REGION Network 8: Concatenadora 2
   RUNG wire#powerrail
      Contact( "EstadosCmpALTA-MTA"._5s4 )
      wire#w1
      { S7_Templates := "SrcType := Int" } NE_Contact(in1 := "CompALTA-MTA".VRealCmp5, in2 := 1)
      wire#w2
      { S7_Templates := "SrcType := Int" } GT_Contact(in1 := "CompALTA-MTA".VRealCmp5, in2 := "CompALTA-MTA".VRealCmp1)
      { S7_Templates := "SrcType := Int" } NE_Contact(in1 := "CompALTA-MTA".VRealCmp1, in2 := 0)
      wire#w3
      Contact( "TV5" )
      wire#w4
      Coil( "Concatenadoras"._5c2 )
   END_RUNG
   RUNG wire#w2
      { S7_Templates := "SrcType := Int" } GT_Contact(in1 := "CompALTA-MTA".VRealCmp5, in2 := "CompALTA-MTA".VRealCmp2)
      { S7_Templates := "SrcType := Int" } NE_Contact(in1 := "CompALTA-MTA".VRealCmp2, in2 := 0)
   END_RUNG wire#w3
   RUNG wire#w2
      { S7_Templates := "SrcType := Int" } GT_Contact(in1 := "CompALTA-MTA".VRealCmp5, in2 := "CompALTA-MTA".VRealCmp3)
      { S7_Templates := "SrcType := Int" } NE_Contact(in1 := "CompALTA-MTA".VRealCmp3, in2 := 0)
   END_RUNG wire#w3
   RUNG wire#w2
      { S7_Templates := "SrcType := Int" } GT_Contact(in1 := "CompALTA-MTA".VRealCmp5, in2 := "CompALTA-MTA".VRealCmp4)
      { S7_Templates := "SrcType := Int" } NE_Contact(in1 := "CompALTA-MTA".VRealCmp4, in2 := 0)
   END_RUNG wire#w3
   RUNG wire#w2
      { S7_Templates := "SrcType := Int" } GT_Contact(in1 := "CompALTA-MTA".VRealCmp5, in2 := "CompALTA-MTA".VRealCmp6)
      { S7_Templates := "SrcType := Int" } NE_Contact(in1 := "CompALTA-MTA".VRealCmp6, in2 := 0)
   END_RUNG wire#w3
   RUNG wire#w1
      Contact( "DB-CompAltaDatos".TON_ParGenMem )
   END_RUNG wire#w4
   RUNG wire#powerrail
      Contact( "EstadosCmpALTA-MTA"._5s6 )
      Contact( "DB-CompAltaDatos".Aut5 )
      Contact( "DB-CompAltaDatos".PanMchCmp5 )
   END_RUNG wire#w4
   // the same network as SCL:
   "Concatenadoras"._5c2 := ("EstadosCmpALTA-MTA"._5s4 AND ((("CompALTA-MTA".VRealCmp5 <> 1) AND ((("CompALTA-MTA".VRealCmp5 > "CompALTA-MTA".VRealCmp1) AND ("CompALTA-MTA".VRealCmp1 <> 0)) OR (("CompALTA-MTA".VRealCmp5 > "CompALTA-MTA".VRealCmp2) AND ("CompALTA-MTA".VRealCmp2 <> 0)) OR (("CompALTA-MTA".VRealCmp5 > "CompALTA-MTA".VRealCmp3) AND ("CompALTA-MTA".VRealCmp3 <> 0)) OR (("CompALTA-MTA".VRealCmp5 > "CompALTA-MTA".VRealCmp4) AND ("CompALTA-MTA".VRealCmp4 <> 0)) OR (("CompALTA-MTA".VRealCmp5 > "CompALTA-MTA".VRealCmp6) AND ("CompALTA-MTA".VRealCmp6 <> 0))) AND "TV5") OR "DB-CompAltaDatos".TON_ParGenMem)) OR ("EstadosCmpALTA-MTA"._5s6 AND "DB-CompAltaDatos".Aut5 AND "DB-CompAltaDatos".PanMchCmp5);
END_REGION

REGION Network 9: Concatenadora 3
   RUNG wire#powerrail
      Contact( "EstadosCmpALTA-MTA"._5s2 )
      Contact( "TsinReq5" )
      wire#w1
      Coil( "Concatenadoras"._5c3 )
   END_RUNG
   RUNG wire#powerrail
      Contact( "EstadosCmpALTA-MTA"._5s10 )
      Contact( "DB-CompAltaDatos".PanMchCmp5 )
   END_RUNG wire#w1
   // the same network as SCL:
   "Concatenadoras"._5c3 := ("EstadosCmpALTA-MTA"._5s2 AND "TsinReq5") OR ("EstadosCmpALTA-MTA"._5s10 AND "DB-CompAltaDatos".PanMchCmp5);
END_REGION

REGION Network 10: Concatenadora 10
   RUNG wire#powerrail
      Contact( "EstadosCmpALTA-MTA"._5s1 )
      I_Contact( "CompALTA-MTA".ReqMch5 )
      wire#w1
      Contact( "DB-CompAltaDatos".Aut5 )
      Coil( "Concatenadoras"._5c10 )
   END_RUNG
   RUNG wire#powerrail
      Contact( "EstadosCmpALTA-MTA"._5s9 )
      I_Contact( "CompALTA-MTA".ReqMch5 )
   END_RUNG wire#w1
   RUNG wire#powerrail
      Contact( "EstadosCmpALTA-MTA"._5s3 )
      I_Contact( "DB-CompAltaDatos".PanMchCmp5 )
   END_RUNG wire#w1
   // the same network as SCL:
   "Concatenadoras"._5c10 := (("EstadosCmpALTA-MTA"._5s1 AND NOT "CompALTA-MTA".ReqMch5) OR ("EstadosCmpALTA-MTA"._5s9 AND NOT "CompALTA-MTA".ReqMch5) OR ("EstadosCmpALTA-MTA"._5s3 AND NOT "DB-CompAltaDatos".PanMchCmp5)) AND "DB-CompAltaDatos".Aut5;
END_REGION

REGION Network 11: Concatenadora 4
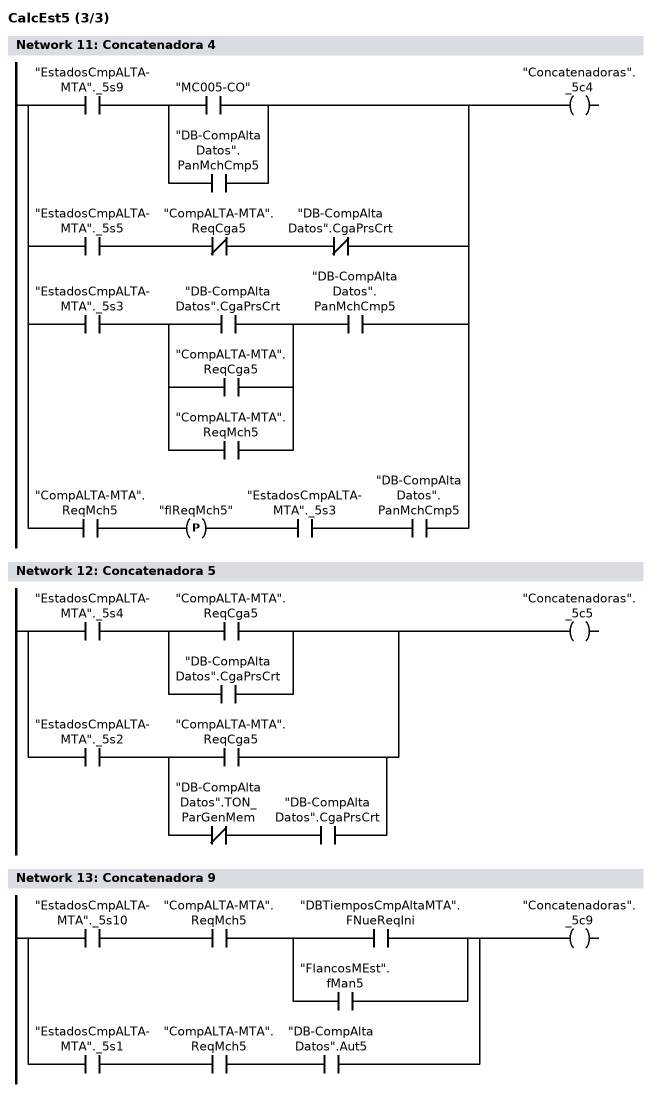
   RUNG wire#powerrail
      Contact( "EstadosCmpALTA-MTA"._5s9 )
      wire#w1
      Contact( "MC005-CO" )
      wire#w2
      Coil( "Concatenadoras"._5c4 )
   END_RUNG
   RUNG wire#w1
      Contact( "DB-CompAltaDatos".PanMchCmp5 )
   END_RUNG wire#w2
   RUNG wire#powerrail
      Contact( "EstadosCmpALTA-MTA"._5s5 )
      I_Contact( "CompALTA-MTA".ReqCga5 )
      I_Contact( "DB-CompAltaDatos".CgaPrsCrt )
   END_RUNG wire#w2
   RUNG wire#powerrail
      Contact( "EstadosCmpALTA-MTA"._5s3 )
      wire#w3
      Contact( "DB-CompAltaDatos".CgaPrsCrt )
      wire#w4
      Contact( "DB-CompAltaDatos".PanMchCmp5 )
   END_RUNG wire#w2
   RUNG wire#w3
      Contact( "CompALTA-MTA".ReqCga5 )
   END_RUNG wire#w4
   RUNG wire#w3
      Contact( "CompALTA-MTA".ReqMch5 )
   END_RUNG wire#w4
   RUNG wire#powerrail
      Contact( "CompALTA-MTA".ReqMch5 )
      P_Trig( "flReqMch5" )
      Contact( "EstadosCmpALTA-MTA"._5s3 )
      Contact( "DB-CompAltaDatos".PanMchCmp5 )
   END_RUNG wire#w2
   // the same network as SCL:
   #_w1 := "CompALTA-MTA".ReqMch5 AND NOT "flReqMch5";   // rising edge
   "flReqMch5" := "CompALTA-MTA".ReqMch5;
   "Concatenadoras"._5c4 := ("EstadosCmpALTA-MTA"._5s9 AND ("MC005-CO" OR "DB-CompAltaDatos".PanMchCmp5)) OR ("EstadosCmpALTA-MTA"._5s5 AND NOT "CompALTA-MTA".ReqCga5 AND NOT "DB-CompAltaDatos".CgaPrsCrt) OR ("EstadosCmpALTA-MTA"._5s3 AND ("DB-CompAltaDatos".CgaPrsCrt OR "CompALTA-MTA".ReqCga5 OR "CompALTA-MTA".ReqMch5) AND "DB-CompAltaDatos".PanMchCmp5) OR (#_w1 AND "EstadosCmpALTA-MTA"._5s3 AND "DB-CompAltaDatos".PanMchCmp5);
END_REGION

REGION Network 12: Concatenadora 5
   RUNG wire#powerrail
      Contact( "EstadosCmpALTA-MTA"._5s4 )
      wire#w1
      Contact( "CompALTA-MTA".ReqCga5 )
      wire#w2
      Coil( "Concatenadoras"._5c5 )
   END_RUNG
   RUNG wire#w1
      Contact( "DB-CompAltaDatos".CgaPrsCrt )
   END_RUNG wire#w2
   RUNG wire#powerrail
      Contact( "EstadosCmpALTA-MTA"._5s2 )
      wire#w3
      Contact( "CompALTA-MTA".ReqCga5 )
   END_RUNG wire#w2
   RUNG wire#w3
      I_Contact( "DB-CompAltaDatos".TON_ParGenMem )
      Contact( "DB-CompAltaDatos".CgaPrsCrt )
   END_RUNG wire#w2
   // the same network as SCL:
   "Concatenadoras"._5c5 := ("EstadosCmpALTA-MTA"._5s4 AND ("CompALTA-MTA".ReqCga5 OR "DB-CompAltaDatos".CgaPrsCrt)) OR ("EstadosCmpALTA-MTA"._5s2 AND ("CompALTA-MTA".ReqCga5 OR (NOT "DB-CompAltaDatos".TON_ParGenMem AND "DB-CompAltaDatos".CgaPrsCrt)));
END_REGION

REGION Network 13: Concatenadora 9
   RUNG wire#powerrail
      Contact( "EstadosCmpALTA-MTA"._5s10 )
      Contact( "CompALTA-MTA".ReqMch5 )
      wire#w1
      Contact( "DBTiemposCmpAltaMTA".FNueReqIni )
      wire#w2
      Coil( "Concatenadoras"._5c9 )
   END_RUNG
   RUNG wire#w1
      Contact( "FlancosMEst".fMan5 )
   END_RUNG wire#w2
   RUNG wire#powerrail
      Contact( "EstadosCmpALTA-MTA"._5s1 )
      Contact( "CompALTA-MTA".ReqMch5 )
      Contact( "DB-CompAltaDatos".Aut5 )
   END_RUNG wire#w2
   // the same network as SCL:
   "Concatenadoras"._5c9 := ("EstadosCmpALTA-MTA"._5s10 AND "CompALTA-MTA".ReqMch5 AND ("DBTiemposCmpAltaMTA".FNueReqIni OR "FlancosMEst".fMan5)) OR ("EstadosCmpALTA-MTA"._5s1 AND "CompALTA-MTA".ReqMch5 AND "DB-CompAltaDatos".Aut5);
END_REGION

REGION Network 14 (STL): Maquina de estados
         CALL  "FC_MAQ_EST_16"
         ( IN0  := %DB127.DBW8,
           IN1  := %DB128.DBW8,
           OUT2 := "ErrPMQ5",
           OUT3 := "ErrCMQ5",
           IO4  := %DB120.DBW8
         );
         NOP   0;
END_REGION

REGION Network 15 (STL): Bloque animación compresor
         CALL  "FC-ANIM-CMP"
         ( IN0  := %DB120.DBW8,
           OUT1 := "CompALTA-MTA".AnimCMP5
         );
         NOP   0;
END_REGION
END_FUNCTION

FUNCTION "CalcEst0" : Void   // FC42, LAD
{ S7_Optimized_Access := 'FALSE' }
VERSION : 0.1
BEGIN

REGION Network 1
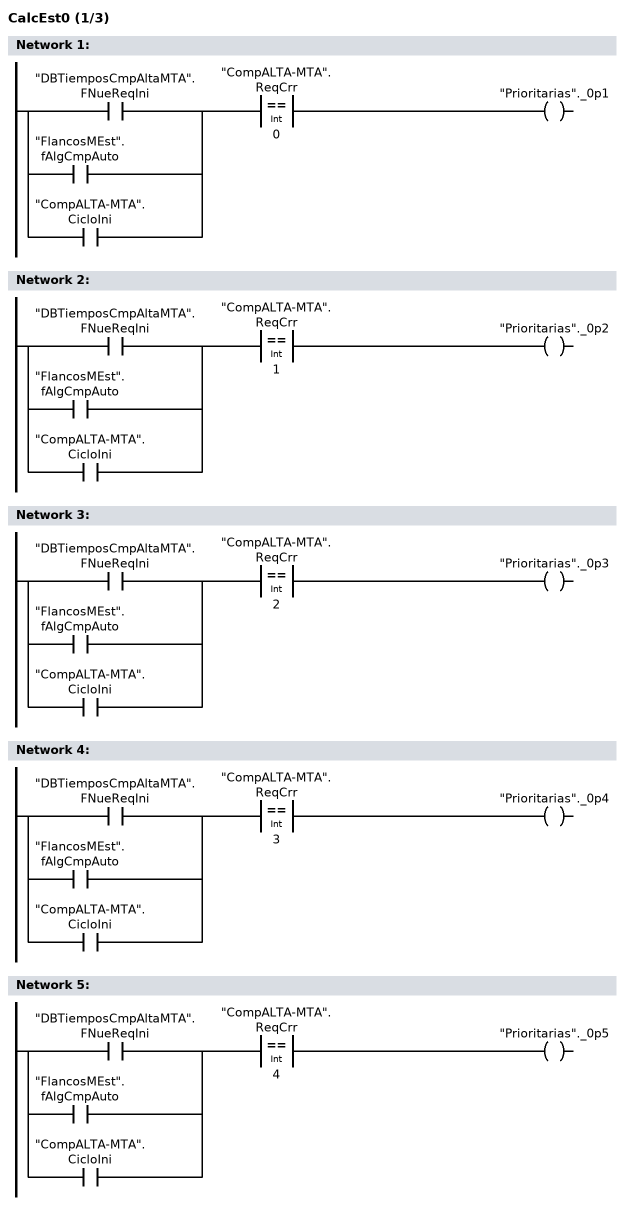
   RUNG wire#powerrail
      Contact( "DBTiemposCmpAltaMTA".FNueReqIni )
      wire#w1
      { S7_Templates := "SrcType := Int" } EQ_Contact(in1 := "CompALTA-MTA".ReqCrr, in2 := 0)
      Coil( "Prioritarias"._0p1 )
   END_RUNG
   RUNG wire#powerrail
      Contact( "FlancosMEst".fAlgCmpAuto )
   END_RUNG wire#w1
   RUNG wire#powerrail
      Contact( "CompALTA-MTA".CicloIni )
   END_RUNG wire#w1
   // the same network as SCL:
   "Prioritarias"._0p1 := ("DBTiemposCmpAltaMTA".FNueReqIni OR "FlancosMEst".fAlgCmpAuto OR "CompALTA-MTA".CicloIni) AND ("CompALTA-MTA".ReqCrr = 0);
END_REGION

REGION Network 2
   RUNG wire#powerrail
      Contact( "DBTiemposCmpAltaMTA".FNueReqIni )
      wire#w1
      { S7_Templates := "SrcType := Int" } EQ_Contact(in1 := "CompALTA-MTA".ReqCrr, in2 := 1)
      Coil( "Prioritarias"._0p2 )
   END_RUNG
   RUNG wire#powerrail
      Contact( "FlancosMEst".fAlgCmpAuto )
   END_RUNG wire#w1
   RUNG wire#powerrail
      Contact( "CompALTA-MTA".CicloIni )
   END_RUNG wire#w1
   // the same network as SCL:
   "Prioritarias"._0p2 := ("DBTiemposCmpAltaMTA".FNueReqIni OR "FlancosMEst".fAlgCmpAuto OR "CompALTA-MTA".CicloIni) AND ("CompALTA-MTA".ReqCrr = 1);
END_REGION

REGION Network 3
   RUNG wire#powerrail
      Contact( "DBTiemposCmpAltaMTA".FNueReqIni )
      wire#w1
      { S7_Templates := "SrcType := Int" } EQ_Contact(in1 := "CompALTA-MTA".ReqCrr, in2 := 2)
      Coil( "Prioritarias"._0p3 )
   END_RUNG
   RUNG wire#powerrail
      Contact( "FlancosMEst".fAlgCmpAuto )
   END_RUNG wire#w1
   RUNG wire#powerrail
      Contact( "CompALTA-MTA".CicloIni )
   END_RUNG wire#w1
   // the same network as SCL:
   "Prioritarias"._0p3 := ("DBTiemposCmpAltaMTA".FNueReqIni OR "FlancosMEst".fAlgCmpAuto OR "CompALTA-MTA".CicloIni) AND ("CompALTA-MTA".ReqCrr = 2);
END_REGION

REGION Network 4
   RUNG wire#powerrail
      Contact( "DBTiemposCmpAltaMTA".FNueReqIni )
      wire#w1
      { S7_Templates := "SrcType := Int" } EQ_Contact(in1 := "CompALTA-MTA".ReqCrr, in2 := 3)
      Coil( "Prioritarias"._0p4 )
   END_RUNG
   RUNG wire#powerrail
      Contact( "FlancosMEst".fAlgCmpAuto )
   END_RUNG wire#w1
   RUNG wire#powerrail
      Contact( "CompALTA-MTA".CicloIni )
   END_RUNG wire#w1
   // the same network as SCL:
   "Prioritarias"._0p4 := ("DBTiemposCmpAltaMTA".FNueReqIni OR "FlancosMEst".fAlgCmpAuto OR "CompALTA-MTA".CicloIni) AND ("CompALTA-MTA".ReqCrr = 3);
END_REGION

REGION Network 5
   RUNG wire#powerrail
      Contact( "DBTiemposCmpAltaMTA".FNueReqIni )
      wire#w1
      { S7_Templates := "SrcType := Int" } EQ_Contact(in1 := "CompALTA-MTA".ReqCrr, in2 := 4)
      Coil( "Prioritarias"._0p5 )
   END_RUNG
   RUNG wire#powerrail
      Contact( "FlancosMEst".fAlgCmpAuto )
   END_RUNG wire#w1
   RUNG wire#powerrail
      Contact( "CompALTA-MTA".CicloIni )
   END_RUNG wire#w1
   // the same network as SCL:
   "Prioritarias"._0p5 := ("DBTiemposCmpAltaMTA".FNueReqIni OR "FlancosMEst".fAlgCmpAuto OR "CompALTA-MTA".CicloIni) AND ("CompALTA-MTA".ReqCrr = 4);
END_REGION

REGION Network 6
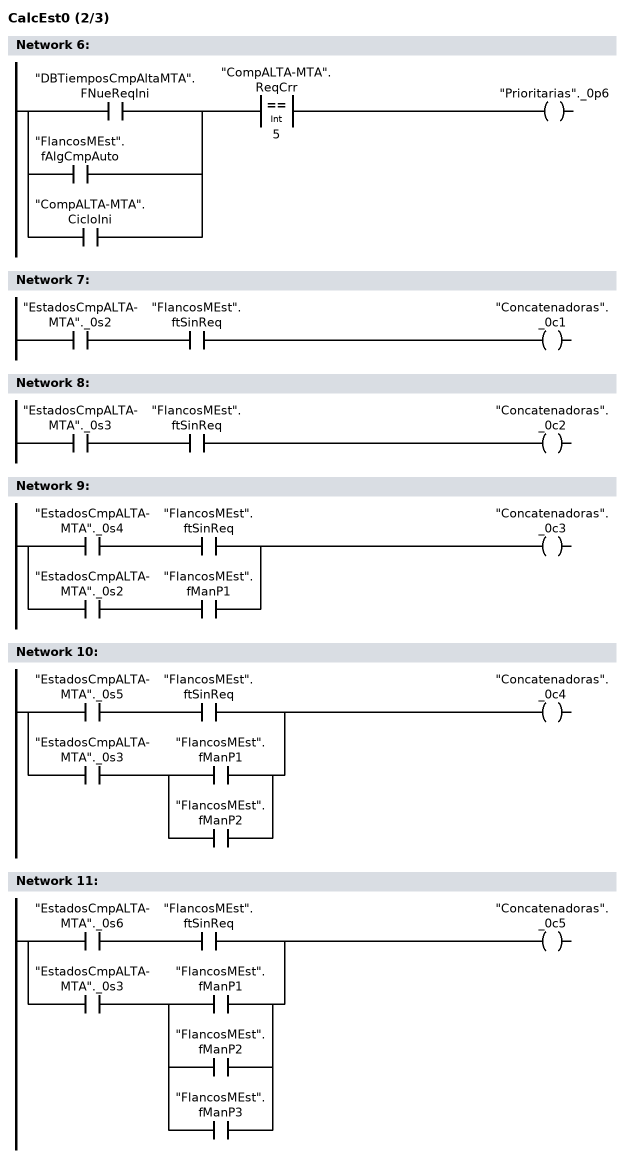
   RUNG wire#powerrail
      Contact( "DBTiemposCmpAltaMTA".FNueReqIni )
      wire#w1
      { S7_Templates := "SrcType := Int" } EQ_Contact(in1 := "CompALTA-MTA".ReqCrr, in2 := 5)
      Coil( "Prioritarias"._0p6 )
   END_RUNG
   RUNG wire#powerrail
      Contact( "FlancosMEst".fAlgCmpAuto )
   END_RUNG wire#w1
   RUNG wire#powerrail
      Contact( "CompALTA-MTA".CicloIni )
   END_RUNG wire#w1
   // the same network as SCL:
   "Prioritarias"._0p6 := ("DBTiemposCmpAltaMTA".FNueReqIni OR "FlancosMEst".fAlgCmpAuto OR "CompALTA-MTA".CicloIni) AND ("CompALTA-MTA".ReqCrr = 5);
END_REGION

REGION Network 7
   RUNG wire#powerrail
      Contact( "EstadosCmpALTA-MTA"._0s2 )
      Contact( "FlancosMEst".ftSinReq )
      Coil( "Concatenadoras"._0c1 )
   END_RUNG
   // the same network as SCL:
   "Concatenadoras"._0c1 := "EstadosCmpALTA-MTA"._0s2 AND "FlancosMEst".ftSinReq;
END_REGION

REGION Network 8
   RUNG wire#powerrail
      Contact( "EstadosCmpALTA-MTA"._0s3 )
      Contact( "FlancosMEst".ftSinReq )
      Coil( "Concatenadoras"._0c2 )
   END_RUNG
   // the same network as SCL:
   "Concatenadoras"._0c2 := "EstadosCmpALTA-MTA"._0s3 AND "FlancosMEst".ftSinReq;
END_REGION

REGION Network 9
   RUNG wire#powerrail
      Contact( "EstadosCmpALTA-MTA"._0s4 )
      Contact( "FlancosMEst".ftSinReq )
      wire#w1
      Coil( "Concatenadoras"._0c3 )
   END_RUNG
   RUNG wire#powerrail
      Contact( "EstadosCmpALTA-MTA"._0s2 )
      Contact( "FlancosMEst".fManP1 )
   END_RUNG wire#w1
   // the same network as SCL:
   "Concatenadoras"._0c3 := ("EstadosCmpALTA-MTA"._0s4 AND "FlancosMEst".ftSinReq) OR ("EstadosCmpALTA-MTA"._0s2 AND "FlancosMEst".fManP1);
END_REGION

REGION Network 10
   RUNG wire#powerrail
      Contact( "EstadosCmpALTA-MTA"._0s5 )
      Contact( "FlancosMEst".ftSinReq )
      wire#w1
      Coil( "Concatenadoras"._0c4 )
   END_RUNG
   RUNG wire#powerrail
      Contact( "EstadosCmpALTA-MTA"._0s3 )
      wire#w2
      Contact( "FlancosMEst".fManP1 )
   END_RUNG wire#w1
   RUNG wire#w2
      Contact( "FlancosMEst".fManP2 )
   END_RUNG wire#w1
   // the same network as SCL:
   "Concatenadoras"._0c4 := ("EstadosCmpALTA-MTA"._0s5 AND "FlancosMEst".ftSinReq) OR ("EstadosCmpALTA-MTA"._0s3 AND ("FlancosMEst".fManP1 OR "FlancosMEst".fManP2));
END_REGION

REGION Network 11
   RUNG wire#powerrail
      Contact( "EstadosCmpALTA-MTA"._0s6 )
      Contact( "FlancosMEst".ftSinReq )
      wire#w1
      Coil( "Concatenadoras"._0c5 )
   END_RUNG
   RUNG wire#powerrail
      Contact( "EstadosCmpALTA-MTA"._0s3 )
      wire#w2
      Contact( "FlancosMEst".fManP1 )
   END_RUNG wire#w1
   RUNG wire#w2
      Contact( "FlancosMEst".fManP2 )
   END_RUNG wire#w1
   RUNG wire#w2
      Contact( "FlancosMEst".fManP3 )
   END_RUNG wire#w1
   // the same network as SCL:
   "Concatenadoras"._0c5 := ("EstadosCmpALTA-MTA"._0s6 AND "FlancosMEst".ftSinReq) OR ("EstadosCmpALTA-MTA"._0s3 AND ("FlancosMEst".fManP1 OR "FlancosMEst".fManP2 OR "FlancosMEst".fManP3));
END_REGION

REGION Network 12
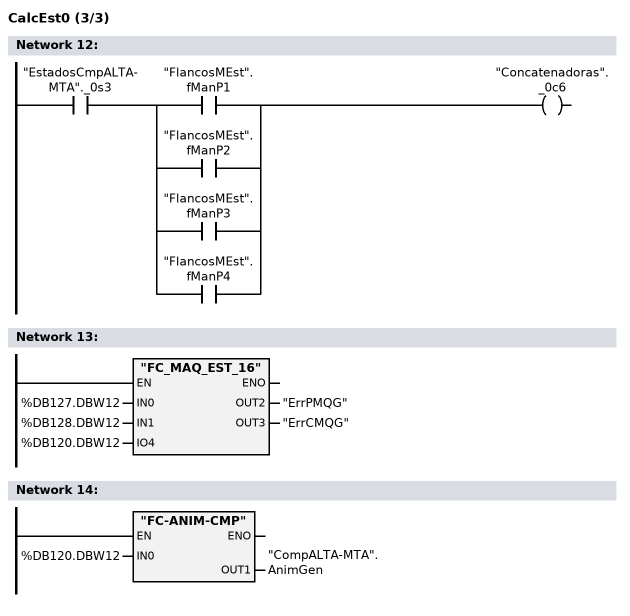
   RUNG wire#powerrail
      Contact( "EstadosCmpALTA-MTA"._0s3 )
      wire#w1
      Contact( "FlancosMEst".fManP1 )
      wire#w2
      Coil( "Concatenadoras"._0c6 )
   END_RUNG
   RUNG wire#w1
      Contact( "FlancosMEst".fManP2 )
   END_RUNG wire#w2
   RUNG wire#w1
      Contact( "FlancosMEst".fManP3 )
   END_RUNG wire#w2
   RUNG wire#w1
      Contact( "FlancosMEst".fManP4 )
   END_RUNG wire#w2
   // the same network as SCL:
   "Concatenadoras"._0c6 := "EstadosCmpALTA-MTA"._0s3 AND ("FlancosMEst".fManP1 OR "FlancosMEst".fManP2 OR "FlancosMEst".fManP3 OR "FlancosMEst".fManP4);
END_REGION

REGION Network 13
   RUNG wire#powerrail
      "FC_MAQ_EST_16"(IN0 := %DB127.DBW12, IN1 := %DB128.DBW12, IO4 := %DB120.DBW12, OUT2 => "ErrPMQG", OUT3 => "ErrCMQG")
   END_RUNG
   // the same network as SCL:
   "FC_MAQ_EST_16"(IN0 := %DB127.DBW12,
                   IN1 := %DB128.DBW12,
                   IO4 := %DB120.DBW12,
                   OUT2 => "ErrPMQG",
                   OUT3 => "ErrCMQG");
END_REGION

REGION Network 14
   RUNG wire#powerrail
      "FC-ANIM-CMP"(IN0 := %DB120.DBW12, OUT1 => "CompALTA-MTA".AnimGen)
   END_RUNG
   // the same network as SCL:
   "FC-ANIM-CMP"(IN0 := %DB120.DBW12, OUT1 => "CompALTA-MTA".AnimGen);
END_REGION
END_FUNCTION

FUNCTION "CorreccReqCmpAlta" : Void   // FC44, LAD
{ S7_Optimized_Access := 'FALSE' }
VERSION : 0.1
BEGIN

REGION Network 1
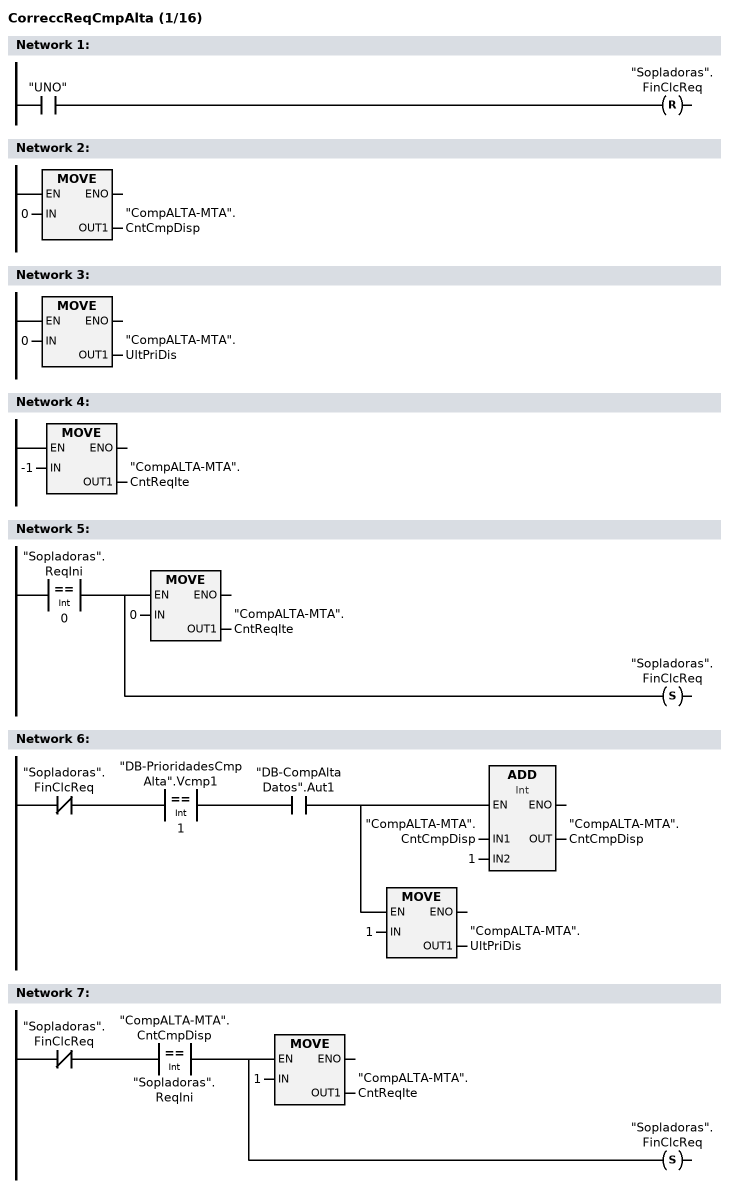
   RUNG wire#powerrail
      Contact( "UNO" )
      R_Coil( "Sopladoras".FinClcReq )
   END_RUNG
   // the same network as SCL:
   IF "UNO" THEN "Sopladoras".FinClcReq := FALSE; END_IF;
END_REGION

REGION Network 2
   RUNG wire#powerrail
      { S7_GenerateENO := "TRUE" } Move(in := 0, out1 => "CompALTA-MTA".CntCmpDisp)
   END_RUNG
   // the same network as SCL:
   "CompALTA-MTA".CntCmpDisp := 0;
END_REGION

REGION Network 3
   RUNG wire#powerrail
      { S7_GenerateENO := "TRUE" } Move(in := 0, out1 => "CompALTA-MTA".UltPriDis)
   END_RUNG
   // the same network as SCL:
   "CompALTA-MTA".UltPriDis := 0;
END_REGION

REGION Network 4
   RUNG wire#powerrail
      { S7_GenerateENO := "TRUE" } Move(in := -1, out1 => "CompALTA-MTA".CntReqIte)
   END_RUNG
   // the same network as SCL:
   "CompALTA-MTA".CntReqIte := -1;
END_REGION

REGION Network 5
   RUNG wire#powerrail
      { S7_Templates := "SrcType := Int" } EQ_Contact(in1 := "Sopladoras".ReqIni, in2 := 0)
      wire#w1
      { S7_GenerateENO := "TRUE" } Move(in := 0, out1 => "CompALTA-MTA".CntReqIte)
   END_RUNG
   RUNG wire#w1
      S_Coil( "Sopladoras".FinClcReq )
   END_RUNG
   // the same network as SCL:
   IF "Sopladoras".ReqIni = 0 THEN
       "CompALTA-MTA".CntReqIte := 0;
       "Sopladoras".FinClcReq := TRUE;
   END_IF;
END_REGION

REGION Network 6
   IF NOT "Sopladoras".FinClcReq AND ("DB-PrioridadesCmpAlta".Vcmp1 = 1) AND "DB-CompAltaDatos".Aut1 THEN
       "CompALTA-MTA".CntCmpDisp := "CompALTA-MTA".CntCmpDisp + 1;
       "CompALTA-MTA".UltPriDis := 1;
   END_IF;
END_REGION

REGION Network 7
   IF NOT "Sopladoras".FinClcReq AND ("CompALTA-MTA".CntCmpDisp = "Sopladoras".ReqIni) THEN
       "CompALTA-MTA".CntReqIte := 1;
       "Sopladoras".FinClcReq := TRUE;
   END_IF;
END_REGION

REGION Network 8
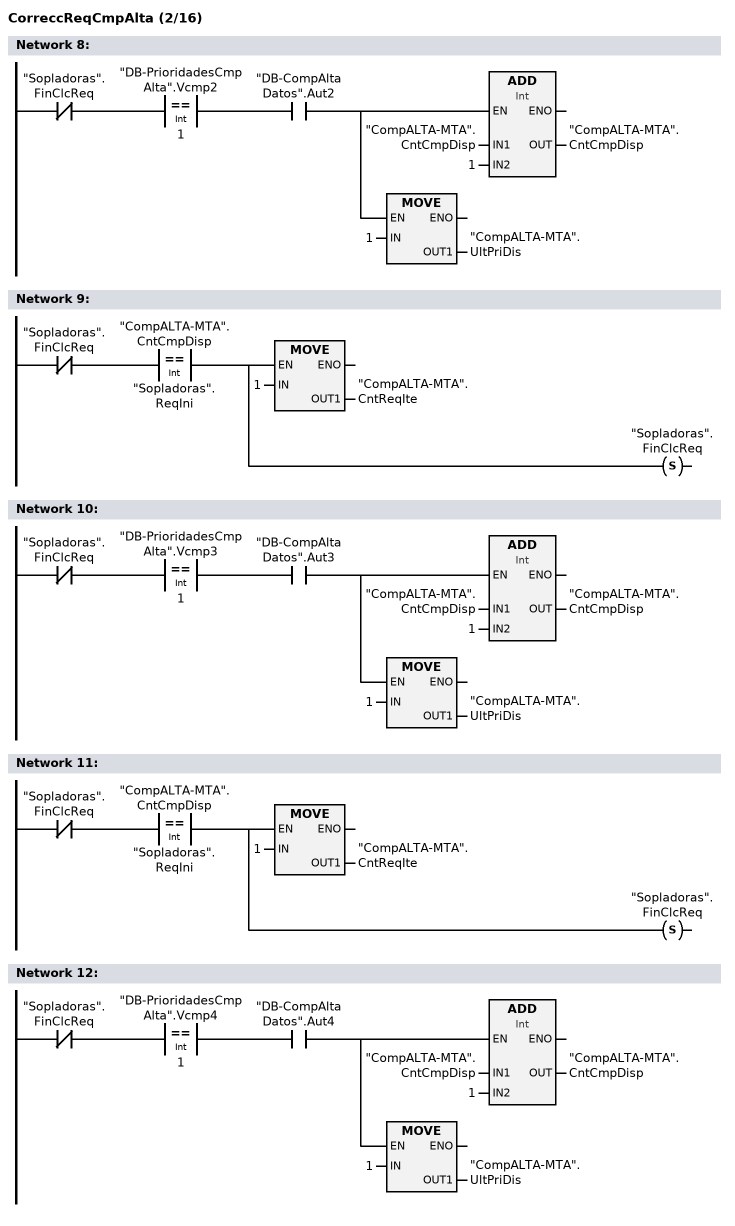
   IF NOT "Sopladoras".FinClcReq AND ("DB-PrioridadesCmpAlta".Vcmp2 = 1) AND "DB-CompAltaDatos".Aut2 THEN
       "CompALTA-MTA".CntCmpDisp := "CompALTA-MTA".CntCmpDisp + 1;
       "CompALTA-MTA".UltPriDis := 1;
   END_IF;
END_REGION

REGION Network 9
   IF NOT "Sopladoras".FinClcReq AND ("CompALTA-MTA".CntCmpDisp = "Sopladoras".ReqIni) THEN
       "CompALTA-MTA".CntReqIte := 1;
       "Sopladoras".FinClcReq := TRUE;
   END_IF;
END_REGION

REGION Network 10
   IF NOT "Sopladoras".FinClcReq AND ("DB-PrioridadesCmpAlta".Vcmp3 = 1) AND "DB-CompAltaDatos".Aut3 THEN
       "CompALTA-MTA".CntCmpDisp := "CompALTA-MTA".CntCmpDisp + 1;
       "CompALTA-MTA".UltPriDis := 1;
   END_IF;
END_REGION

REGION Network 11
   IF NOT "Sopladoras".FinClcReq AND ("CompALTA-MTA".CntCmpDisp = "Sopladoras".ReqIni) THEN
       "CompALTA-MTA".CntReqIte := 1;
       "Sopladoras".FinClcReq := TRUE;
   END_IF;
END_REGION

REGION Network 12
   IF NOT "Sopladoras".FinClcReq AND ("DB-PrioridadesCmpAlta".Vcmp4 = 1) AND "DB-CompAltaDatos".Aut4 THEN
       "CompALTA-MTA".CntCmpDisp := "CompALTA-MTA".CntCmpDisp + 1;
       "CompALTA-MTA".UltPriDis := 1;
   END_IF;
END_REGION

REGION Network 13
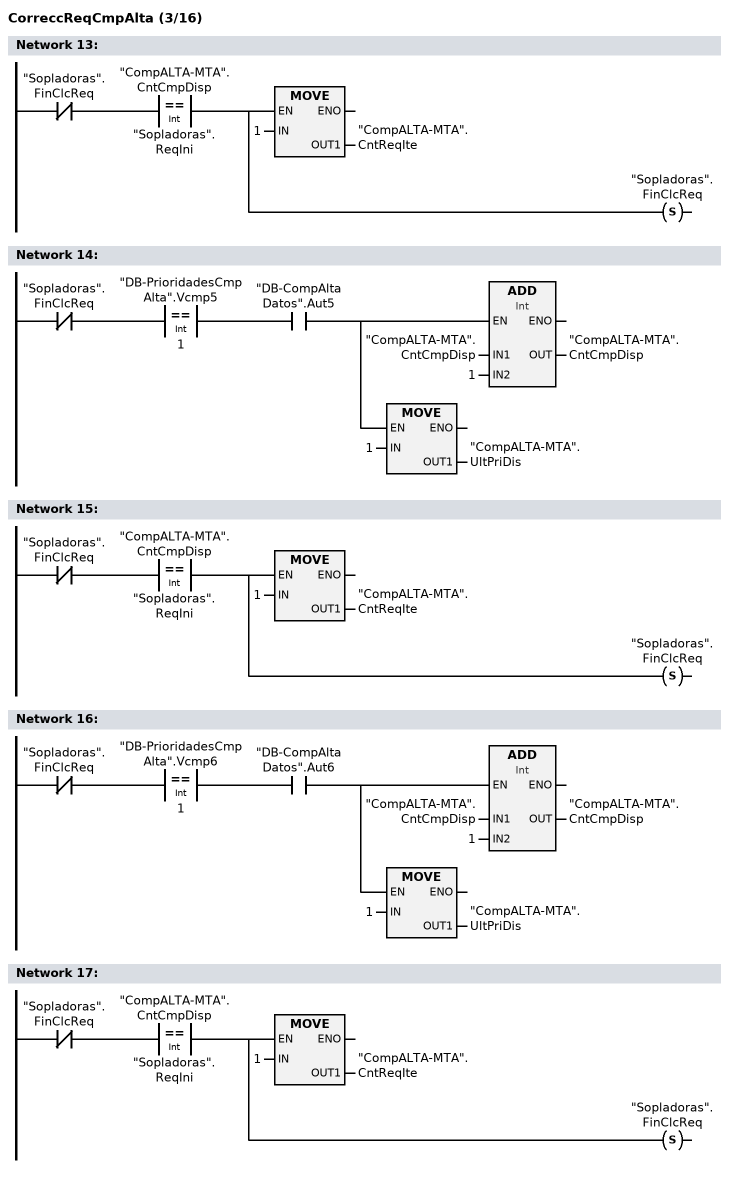
   IF NOT "Sopladoras".FinClcReq AND ("CompALTA-MTA".CntCmpDisp = "Sopladoras".ReqIni) THEN
       "CompALTA-MTA".CntReqIte := 1;
       "Sopladoras".FinClcReq := TRUE;
   END_IF;
END_REGION

REGION Network 14
   IF NOT "Sopladoras".FinClcReq AND ("DB-PrioridadesCmpAlta".Vcmp5 = 1) AND "DB-CompAltaDatos".Aut5 THEN
       "CompALTA-MTA".CntCmpDisp := "CompALTA-MTA".CntCmpDisp + 1;
       "CompALTA-MTA".UltPriDis := 1;
   END_IF;
END_REGION

REGION Network 15
   IF NOT "Sopladoras".FinClcReq AND ("CompALTA-MTA".CntCmpDisp = "Sopladoras".ReqIni) THEN
       "CompALTA-MTA".CntReqIte := 1;
       "Sopladoras".FinClcReq := TRUE;
   END_IF;
END_REGION

REGION Network 16
   RUNG wire#powerrail
      I_Contact( "Sopladoras".FinClcReq )
      { S7_Templates := "SrcType := Int" } EQ_Contact(in1 := "DB-PrioridadesCmpAlta".Vcmp6, in2 := 1)
      Contact( "DB-CompAltaDatos".Aut6 )
      wire#w1
      { S7_Templates := "SrcType := Int"; S7_GenerateENO := "TRUE" } Add(in1 := "CompALTA-MTA".CntCmpDisp, in2 := 1, out => "CompALTA-MTA".CntCmpDisp)
   END_RUNG
   RUNG wire#w1
      { S7_GenerateENO := "TRUE" } Move(in := 1, out1 => "CompALTA-MTA".UltPriDis)
   END_RUNG
   // the same network as SCL:
   IF NOT "Sopladoras".FinClcReq AND ("DB-PrioridadesCmpAlta".Vcmp6 = 1) AND "DB-CompAltaDatos".Aut6 THEN
       "CompALTA-MTA".CntCmpDisp := "CompALTA-MTA".CntCmpDisp + 1;
       "CompALTA-MTA".UltPriDis := 1;
   END_IF;
END_REGION

REGION Network 17
   RUNG wire#powerrail
      I_Contact( "Sopladoras".FinClcReq )
      { S7_Templates := "SrcType := Int" } EQ_Contact(in1 := "CompALTA-MTA".CntCmpDisp, in2 := "Sopladoras".ReqIni)
      wire#w1
      { S7_GenerateENO := "TRUE" } Move(in := 1, out1 => "CompALTA-MTA".CntReqIte)
   END_RUNG
   RUNG wire#w1
      S_Coil( "Sopladoras".FinClcReq )
   END_RUNG
   // the same network as SCL:
   IF NOT "Sopladoras".FinClcReq AND ("CompALTA-MTA".CntCmpDisp = "Sopladoras".ReqIni) THEN
       "CompALTA-MTA".CntReqIte := 1;
       "Sopladoras".FinClcReq := TRUE;
   END_IF;
END_REGION

REGION Network 18
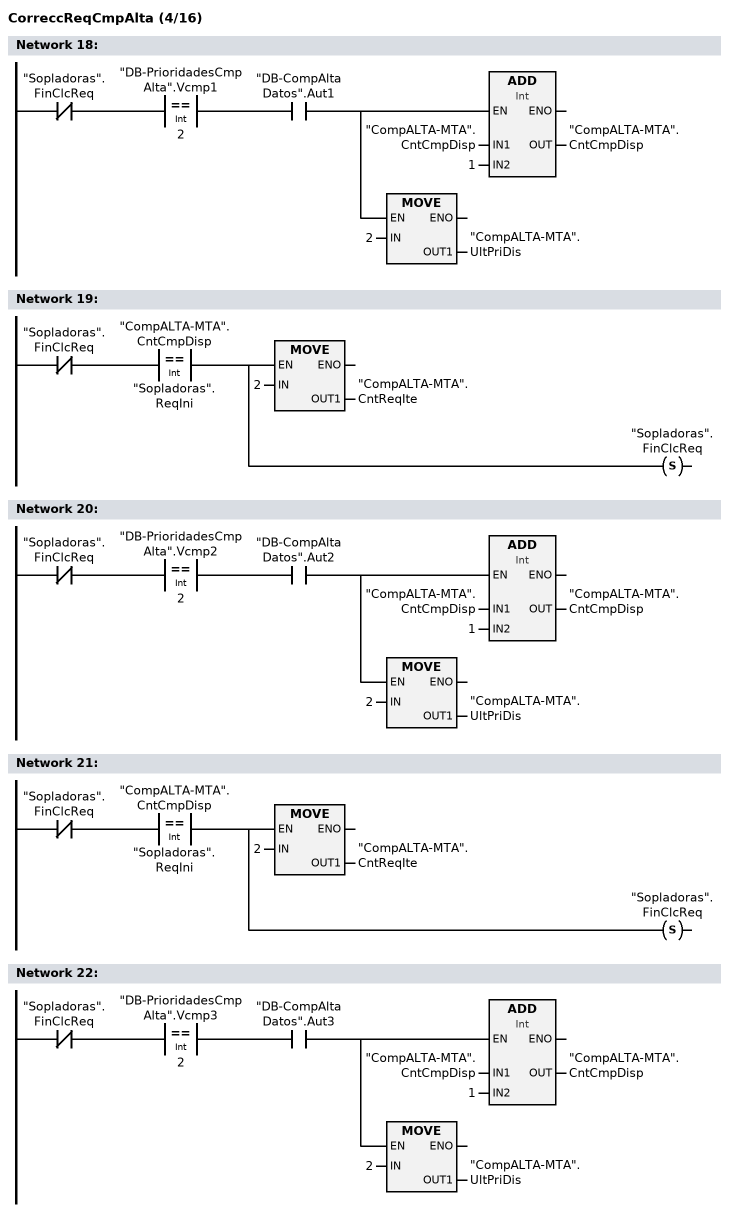
   IF NOT "Sopladoras".FinClcReq AND ("DB-PrioridadesCmpAlta".Vcmp1 = 2) AND "DB-CompAltaDatos".Aut1 THEN
       "CompALTA-MTA".CntCmpDisp := "CompALTA-MTA".CntCmpDisp + 1;
       "CompALTA-MTA".UltPriDis := 2;
   END_IF;
END_REGION

REGION Network 19
   IF NOT "Sopladoras".FinClcReq AND ("CompALTA-MTA".CntCmpDisp = "Sopladoras".ReqIni) THEN
       "CompALTA-MTA".CntReqIte := 2;
       "Sopladoras".FinClcReq := TRUE;
   END_IF;
END_REGION

REGION Network 20
   IF NOT "Sopladoras".FinClcReq AND ("DB-PrioridadesCmpAlta".Vcmp2 = 2) AND "DB-CompAltaDatos".Aut2 THEN
       "CompALTA-MTA".CntCmpDisp := "CompALTA-MTA".CntCmpDisp + 1;
       "CompALTA-MTA".UltPriDis := 2;
   END_IF;
END_REGION

REGION Network 21
   IF NOT "Sopladoras".FinClcReq AND ("CompALTA-MTA".CntCmpDisp = "Sopladoras".ReqIni) THEN
       "CompALTA-MTA".CntReqIte := 2;
       "Sopladoras".FinClcReq := TRUE;
   END_IF;
END_REGION

REGION Network 22
   IF NOT "Sopladoras".FinClcReq AND ("DB-PrioridadesCmpAlta".Vcmp3 = 2) AND "DB-CompAltaDatos".Aut3 THEN
       "CompALTA-MTA".CntCmpDisp := "CompALTA-MTA".CntCmpDisp + 1;
       "CompALTA-MTA".UltPriDis := 2;
   END_IF;
END_REGION

REGION Network 23
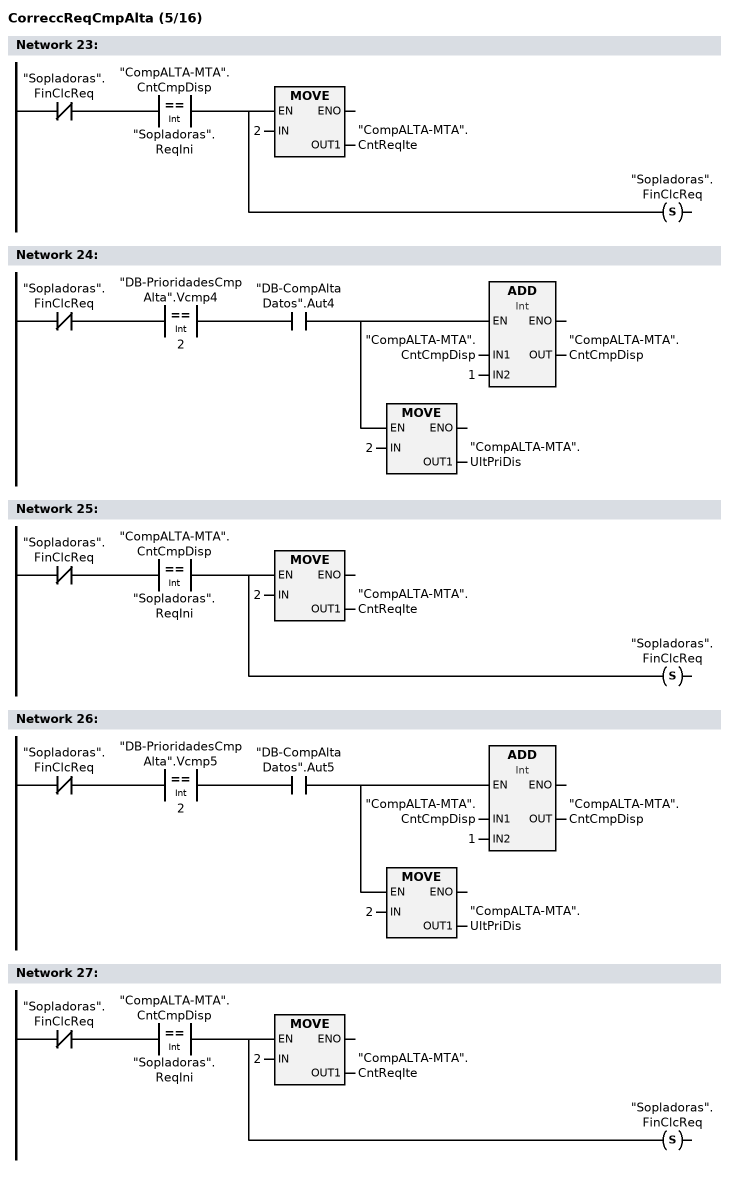
   IF NOT "Sopladoras".FinClcReq AND ("CompALTA-MTA".CntCmpDisp = "Sopladoras".ReqIni) THEN
       "CompALTA-MTA".CntReqIte := 2;
       "Sopladoras".FinClcReq := TRUE;
   END_IF;
END_REGION

REGION Network 24
   IF NOT "Sopladoras".FinClcReq AND ("DB-PrioridadesCmpAlta".Vcmp4 = 2) AND "DB-CompAltaDatos".Aut4 THEN
       "CompALTA-MTA".CntCmpDisp := "CompALTA-MTA".CntCmpDisp + 1;
       "CompALTA-MTA".UltPriDis := 2;
   END_IF;
END_REGION

REGION Network 25
   IF NOT "Sopladoras".FinClcReq AND ("CompALTA-MTA".CntCmpDisp = "Sopladoras".ReqIni) THEN
       "CompALTA-MTA".CntReqIte := 2;
       "Sopladoras".FinClcReq := TRUE;
   END_IF;
END_REGION

REGION Network 26
   IF NOT "Sopladoras".FinClcReq AND ("DB-PrioridadesCmpAlta".Vcmp5 = 2) AND "DB-CompAltaDatos".Aut5 THEN
       "CompALTA-MTA".CntCmpDisp := "CompALTA-MTA".CntCmpDisp + 1;
       "CompALTA-MTA".UltPriDis := 2;
   END_IF;
END_REGION

REGION Network 27
   IF NOT "Sopladoras".FinClcReq AND ("CompALTA-MTA".CntCmpDisp = "Sopladoras".ReqIni) THEN
       "CompALTA-MTA".CntReqIte := 2;
       "Sopladoras".FinClcReq := TRUE;
   END_IF;
END_REGION

REGION Network 28
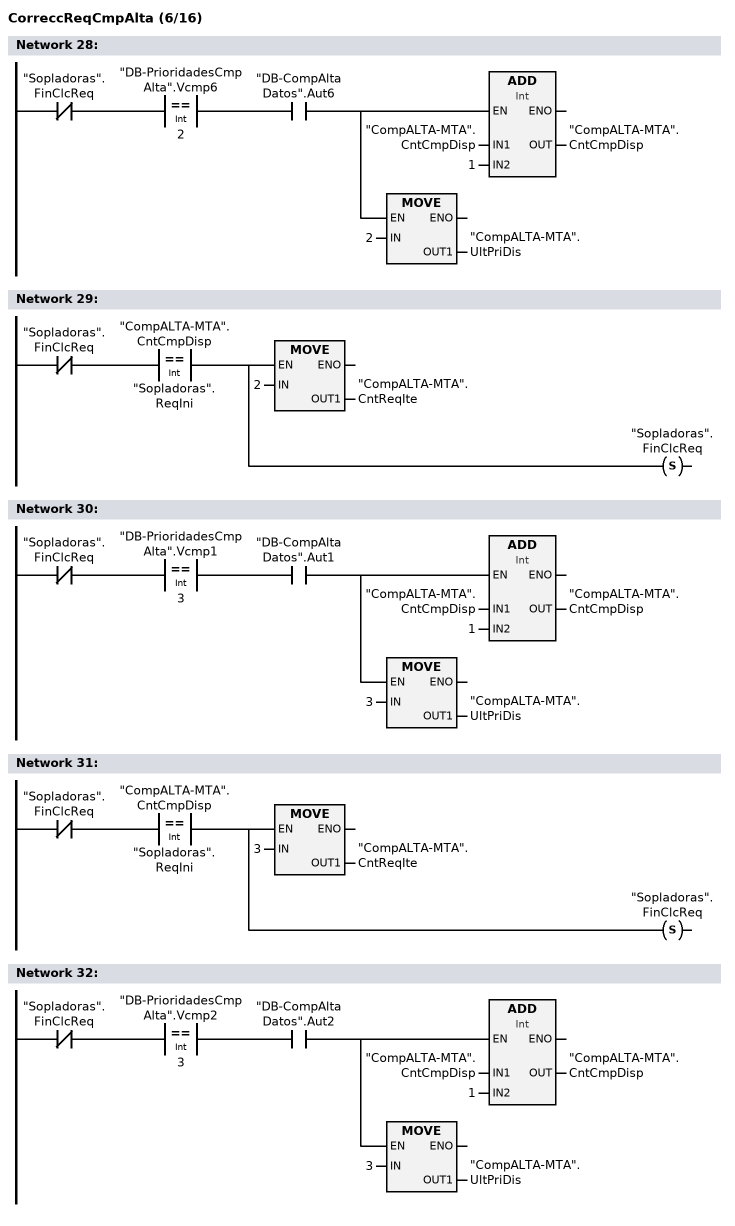
   RUNG wire#powerrail
      I_Contact( "Sopladoras".FinClcReq )
      { S7_Templates := "SrcType := Int" } EQ_Contact(in1 := "DB-PrioridadesCmpAlta".Vcmp6, in2 := 2)
      Contact( "DB-CompAltaDatos".Aut6 )
      wire#w1
      { S7_Templates := "SrcType := Int"; S7_GenerateENO := "TRUE" } Add(in1 := "CompALTA-MTA".CntCmpDisp, in2 := 1, out => "CompALTA-MTA".CntCmpDisp)
   END_RUNG
   RUNG wire#w1
      { S7_GenerateENO := "TRUE" } Move(in := 2, out1 => "CompALTA-MTA".UltPriDis)
   END_RUNG
   // the same network as SCL:
   IF NOT "Sopladoras".FinClcReq AND ("DB-PrioridadesCmpAlta".Vcmp6 = 2) AND "DB-CompAltaDatos".Aut6 THEN
       "CompALTA-MTA".CntCmpDisp := "CompALTA-MTA".CntCmpDisp + 1;
       "CompALTA-MTA".UltPriDis := 2;
   END_IF;
END_REGION

REGION Network 29
   RUNG wire#powerrail
      I_Contact( "Sopladoras".FinClcReq )
      { S7_Templates := "SrcType := Int" } EQ_Contact(in1 := "CompALTA-MTA".CntCmpDisp, in2 := "Sopladoras".ReqIni)
      wire#w1
      { S7_GenerateENO := "TRUE" } Move(in := 2, out1 => "CompALTA-MTA".CntReqIte)
   END_RUNG
   RUNG wire#w1
      S_Coil( "Sopladoras".FinClcReq )
   END_RUNG
   // the same network as SCL:
   IF NOT "Sopladoras".FinClcReq AND ("CompALTA-MTA".CntCmpDisp = "Sopladoras".ReqIni) THEN
       "CompALTA-MTA".CntReqIte := 2;
       "Sopladoras".FinClcReq := TRUE;
   END_IF;
END_REGION

REGION Network 30
   IF NOT "Sopladoras".FinClcReq AND ("DB-PrioridadesCmpAlta".Vcmp1 = 3) AND "DB-CompAltaDatos".Aut1 THEN
       "CompALTA-MTA".CntCmpDisp := "CompALTA-MTA".CntCmpDisp + 1;
       "CompALTA-MTA".UltPriDis := 3;
   END_IF;
END_REGION

REGION Network 31
   IF NOT "Sopladoras".FinClcReq AND ("CompALTA-MTA".CntCmpDisp = "Sopladoras".ReqIni) THEN
       "CompALTA-MTA".CntReqIte := 3;
       "Sopladoras".FinClcReq := TRUE;
   END_IF;
END_REGION

REGION Network 32
   IF NOT "Sopladoras".FinClcReq AND ("DB-PrioridadesCmpAlta".Vcmp2 = 3) AND "DB-CompAltaDatos".Aut2 THEN
       "CompALTA-MTA".CntCmpDisp := "CompALTA-MTA".CntCmpDisp + 1;
       "CompALTA-MTA".UltPriDis := 3;
   END_IF;
END_REGION

REGION Network 33
